// TIA Portal project "uppgift2IndustriellIT" (V18) (continued)
REGION Network 9: if x or y arm is moving for hmi
   RUNG wire#powerrail
      Contact( "InputsDB".Crane.RunArmX )
      { S7_Templates := "SrcType := Int" } NE_Contact(in1 := "Crane Current X Position", in2 := "OutputsDB".CraneOutput.XScalex)
      Coil( "InputsDB".XisMoving )
   END_RUNG
   RUNG wire#powerrail
      Contact( "InputsDB".Crane.RunArmY )
      { S7_Templates := "SrcType := Int" } NE_Contact(in1 := "Crane Current Z Position", in2 := "OutputsDB".CraneOutput.YScalex)
      Coil( "InputsDB".YisMoving )
   END_RUNG
   // the same network as SCL:
   "InputsDB".XisMoving := "InputsDB".Crane.RunArmX AND ("Crane Current X Position" <> "OutputsDB".CraneOutput.XScalex);
   "InputsDB".YisMoving := "InputsDB".Crane.RunArmY AND ("Crane Current Z Position" <> "OutputsDB".CraneOutput.YScalex);
END_REGION
END_FUNCTION

FUNCTION "Outputs" : Void   // FC4, LAD
{ S7_Optimized_Access := 'TRUE' }
VERSION : 0.1
   VAR_TEMP   // added for the SCL form of the ladder/FBD networks
      _w1 : Bool;
      _w2 : Bool;
      _w3 : Bool;
      _w4 : Bool;
   END_VAR
BEGIN

REGION Network 1: Convert MM to raw sensor value which is 27648
   // Calling for example "OutputsDB".CraneOutput.Xmm" with a value from 0-10500mm is going to make the crane move.
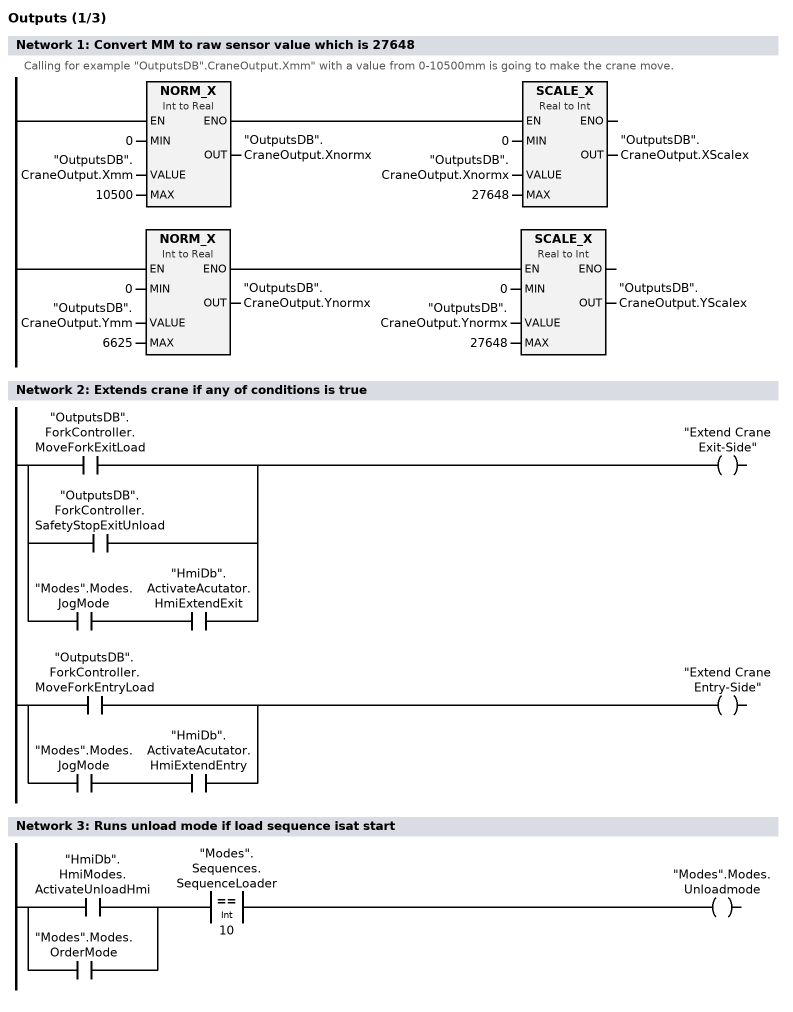
   RUNG wire#powerrail
      { S7_Templates := "[SrcType := Int, DestType := Real]" } Normalize(min := 0, value := "OutputsDB".CraneOutput.Xmm, max := 10500, out => "OutputsDB".CraneOutput.Xnormx)
      { S7_Templates := "[SrcType := Real, DestType := Int]" } Scale(min := 0, value := "OutputsDB".CraneOutput.Xnormx, max := 27648, out => "OutputsDB".CraneOutput.XScalex)
   END_RUNG
   RUNG wire#powerrail
      { S7_Templates := "[SrcType := Int, DestType := Real]" } Normalize(min := 0, value := "OutputsDB".CraneOutput.Ymm, max := 6625, out => "OutputsDB".CraneOutput.Ynormx)
      { S7_Templates := "[SrcType := Real, DestType := Int]" } Scale(min := 0, value := "OutputsDB".CraneOutput.Ynormx, max := 27648, out => "OutputsDB".CraneOutput.YScalex)
   END_RUNG
   // the same network as SCL:
   "OutputsDB".CraneOutput.Xnormx := NORM_X(MIN := 0, VALUE := "OutputsDB".CraneOutput.Xmm, MAX := 10500);
   "OutputsDB".CraneOutput.XScalex := SCALE_X(MIN := 0, VALUE := "OutputsDB".CraneOutput.Xnormx, MAX := 27648);
   "OutputsDB".CraneOutput.Ynormx := NORM_X(MIN := 0, VALUE := "OutputsDB".CraneOutput.Ymm, MAX := 6625);
   "OutputsDB".CraneOutput.YScalex := SCALE_X(MIN := 0, VALUE := "OutputsDB".CraneOutput.Ynormx, MAX := 27648);
END_REGION

REGION Network 2: Extends crane if any of conditions is true
   RUNG wire#powerrail
      Contact( "OutputsDB".ForkController.MoveForkExitLoad )
      wire#w1
      Coil( "Extend Crane Exit-Side" )
   END_RUNG
   RUNG wire#powerrail
      Contact( "OutputsDB".ForkController.SafetyStopExitUnload )
   END_RUNG wire#w1
   RUNG wire#powerrail
      Contact( "Modes".Modes.JogMode )
      Contact( "HmiDb".ActivateAcutator.HmiExtendExit )
   END_RUNG wire#w1
   RUNG wire#powerrail
      Contact( "OutputsDB".ForkController.MoveForkEntryLoad )
      wire#w2
      Coil( "Extend Crane Entry-Side" )
   END_RUNG
   RUNG wire#powerrail
      Contact( "Modes".Modes.JogMode )
      Contact( "HmiDb".ActivateAcutator.HmiExtendEntry )
   END_RUNG wire#w2
   // the same network as SCL:
   "Extend Crane Exit-Side" := "OutputsDB".ForkController.MoveForkExitLoad OR "OutputsDB".ForkController.SafetyStopExitUnload OR ("Modes".Modes.JogMode AND "HmiDb".ActivateAcutator.HmiExtendExit);
   "Extend Crane Entry-Side" := "OutputsDB".ForkController.MoveForkEntryLoad OR ("Modes".Modes.JogMode AND "HmiDb".ActivateAcutator.HmiExtendEntry);
END_REGION

REGION Network 3: Runs unload mode if load sequence isat start
   RUNG wire#powerrail
      Contact( "HmiDb".HmiModes.ActivateUnloadHmi )
      wire#w1
      { S7_Templates := "SrcType := Int" } EQ_Contact(in1 := "Modes".Sequences.SequenceLoader, in2 := 10)
      Coil( "Modes".Modes.Unloadmode )
   END_RUNG
   RUNG wire#powerrail
      Contact( "Modes".Modes.OrderMode )
   END_RUNG wire#w1
   // the same network as SCL:
   "Modes".Modes.Unloadmode := ("HmiDb".HmiModes.ActivateUnloadHmi OR "Modes".Modes.OrderMode) AND ("Modes".Sequences.SequenceLoader = 10);
END_REGION

REGION Network 4: Sets the conveyor speed
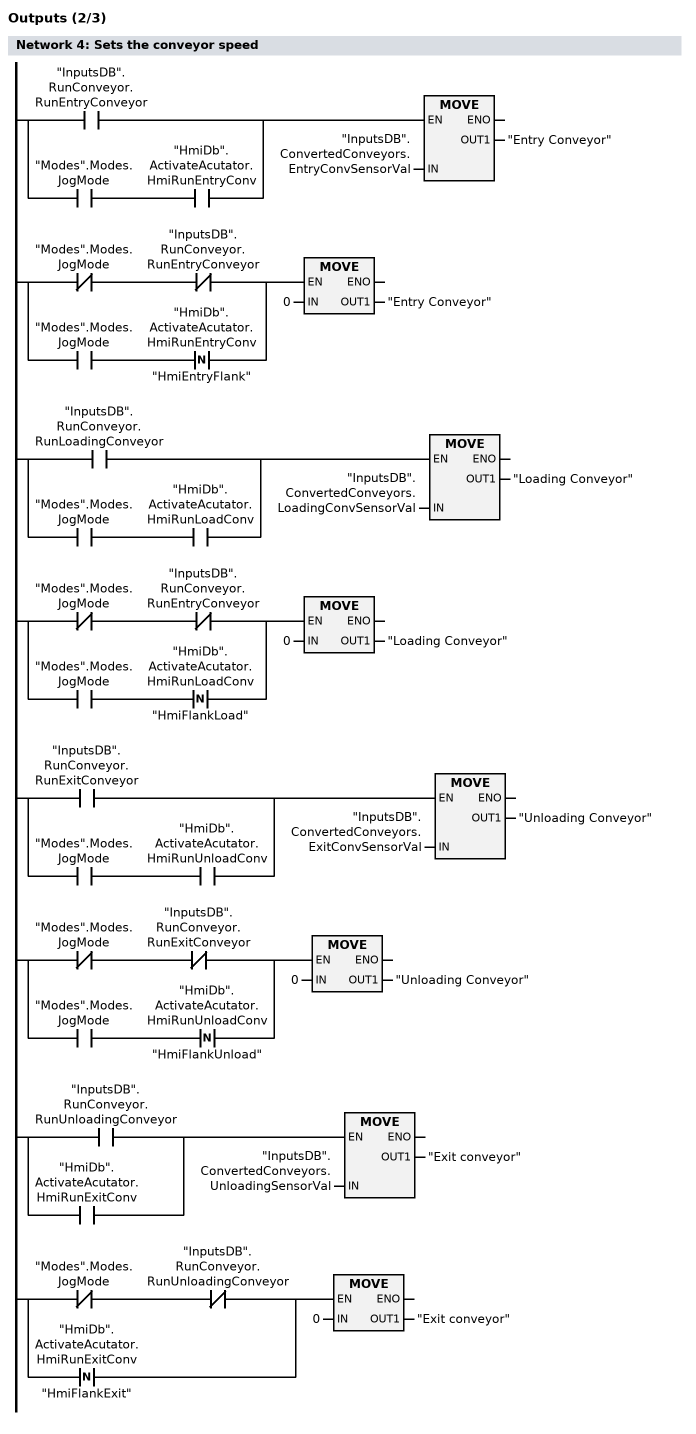
   RUNG wire#powerrail
      Contact( "InputsDB".RunConveyor.RunEntryConveyor )
      wire#w1
      Move(in := "InputsDB".ConvertedConveyors.EntryConvSensorVal, out1 => "Entry Conveyor")
   END_RUNG
   RUNG wire#powerrail
      Contact( "Modes".Modes.JogMode )
      Contact( "HmiDb".ActivateAcutator.HmiRunEntryConv )
   END_RUNG wire#w1
   RUNG wire#powerrail
      I_Contact( "Modes".Modes.JogMode )
      I_Contact( "InputsDB".RunConveyor.RunEntryConveyor )
      wire#w2
      Move(in := 0, out1 => "Entry Conveyor")
   END_RUNG
   RUNG wire#powerrail
      Contact( "Modes".Modes.JogMode )
      N_Contact(operand := "HmiDb".ActivateAcutator.HmiRunEntryConv, bit := "HmiEntryFlank")
   END_RUNG wire#w2
   RUNG wire#powerrail
      Contact( "InputsDB".RunConveyor.RunLoadingConveyor )
      wire#w3
      Move(in := "InputsDB".ConvertedConveyors.LoadingConvSensorVal, out1 => "Loading Conveyor")
   END_RUNG
   RUNG wire#powerrail
      Contact( "Modes".Modes.JogMode )
      Contact( "HmiDb".ActivateAcutator.HmiRunLoadConv )
   END_RUNG wire#w3
   RUNG wire#powerrail
      I_Contact( "Modes".Modes.JogMode )
      I_Contact( "InputsDB".RunConveyor.RunEntryConveyor )
      wire#w4
      Move(in := 0, out1 => "Loading Conveyor")
   END_RUNG
   RUNG wire#powerrail
      Contact( "Modes".Modes.JogMode )
      N_Contact(operand := "HmiDb".ActivateAcutator.HmiRunLoadConv, bit := "HmiFlankLoad")
   END_RUNG wire#w4
   RUNG wire#powerrail
      Contact( "InputsDB".RunConveyor.RunExitConveyor )
      wire#w5
      Move(in := "InputsDB".ConvertedConveyors.ExitConvSensorVal, out1 => "Unloading Conveyor")
   END_RUNG
   RUNG wire#powerrail
      Contact( "Modes".Modes.JogMode )
      Contact( "HmiDb".ActivateAcutator.HmiRunUnloadConv )
   END_RUNG wire#w5
   RUNG wire#powerrail
      I_Contact( "Modes".Modes.JogMode )
      I_Contact( "InputsDB".RunConveyor.RunExitConveyor )
      wire#w6
      Move(in := 0, out1 => "Unloading Conveyor")
   END_RUNG
   RUNG wire#powerrail
      Contact( "Modes".Modes.JogMode )
      N_Contact(operand := "HmiDb".ActivateAcutator.HmiRunUnloadConv, bit := "HmiFlankUnload")
   END_RUNG wire#w6
   RUNG wire#powerrail
      Contact( "InputsDB".RunConveyor.RunUnloadingConveyor )
      wire#w7
      Move(in := "InputsDB".ConvertedConveyors.UnloadingSensorVal, out1 => "Exit conveyor")
   END_RUNG
   RUNG wire#powerrail
      Contact( "HmiDb".ActivateAcutator.HmiRunExitConv )
   END_RUNG wire#w7
   RUNG wire#powerrail
      I_Contact( "Modes".Modes.JogMode )
      I_Contact( "InputsDB".RunConveyor.RunUnloadingConveyor )
      wire#w8
      Move(in := 0, out1 => "Exit conveyor")
   END_RUNG
   RUNG wire#powerrail
      N_Contact(operand := "HmiDb".ActivateAcutator.HmiRunExitConv, bit := "HmiFlankExit")
   END_RUNG wire#w8
   // the same network as SCL:
   IF "InputsDB".RunConveyor.RunEntryConveyor OR ("Modes".Modes.JogMode AND "HmiDb".ActivateAcutator.HmiRunEntryConv) THEN
       "Entry Conveyor" := "InputsDB".ConvertedConveyors.EntryConvSensorVal;
   END_IF;
   #_w1 := "Modes".Modes.JogMode AND NOT "HmiDb".ActivateAcutator.HmiRunEntryConv AND "HmiEntryFlank";   // falling edge of "HmiDb".ActivateAcutator.HmiRunEntryConv
   "HmiEntryFlank" := "HmiDb".ActivateAcutator.HmiRunEntryConv;
   IF (NOT "Modes".Modes.JogMode AND NOT "InputsDB".RunConveyor.RunEntryConveyor) OR #_w1 THEN
       "Entry Conveyor" := 0;
   END_IF;
   IF "InputsDB".RunConveyor.RunLoadingConveyor OR ("Modes".Modes.JogMode AND "HmiDb".ActivateAcutator.HmiRunLoadConv) THEN
       "Loading Conveyor" := "InputsDB".ConvertedConveyors.LoadingConvSensorVal;
   END_IF;
   #_w2 := "Modes".Modes.JogMode AND NOT "HmiDb".ActivateAcutator.HmiRunLoadConv AND "HmiFlankLoad";   // falling edge of "HmiDb".ActivateAcutator.HmiRunLoadConv
   "HmiFlankLoad" := "HmiDb".ActivateAcutator.HmiRunLoadConv;
   IF (NOT "Modes".Modes.JogMode AND NOT "InputsDB".RunConveyor.RunEntryConveyor) OR #_w2 THEN
       "Loading Conveyor" := 0;
   END_IF;
   IF "InputsDB".RunConveyor.RunExitConveyor OR ("Modes".Modes.JogMode AND "HmiDb".ActivateAcutator.HmiRunUnloadConv) THEN
       "Unloading Conveyor" := "InputsDB".ConvertedConveyors.ExitConvSensorVal;
   END_IF;
   #_w3 := "Modes".Modes.JogMode AND NOT "HmiDb".ActivateAcutator.HmiRunUnloadConv AND "HmiFlankUnload";   // falling edge of "HmiDb".ActivateAcutator.HmiRunUnloadConv
   "HmiFlankUnload" := "HmiDb".ActivateAcutator.HmiRunUnloadConv;
   IF (NOT "Modes".Modes.JogMode AND NOT "InputsDB".RunConveyor.RunExitConveyor) OR #_w3 THEN
       "Unloading Conveyor" := 0;
   END_IF;
   IF "InputsDB".RunConveyor.RunUnloadingConveyor OR "HmiDb".ActivateAcutator.HmiRunExitConv THEN
       "Exit conveyor" := "InputsDB".ConvertedConveyors.UnloadingSensorVal;
   END_IF;
   #_w4 := NOT "HmiDb".ActivateAcutator.HmiRunExitConv AND "HmiFlankExit";   // falling edge of "HmiDb".ActivateAcutator.HmiRunExitConv
   "HmiFlankExit" := "HmiDb".ActivateAcutator.HmiRunExitConv;
   IF (NOT "Modes".Modes.JogMode AND NOT "InputsDB".RunConveyor.RunUnloadingConveyor) OR #_w4 THEN
       "Exit conveyor" := 0;
   END_IF;
END_REGION

REGION Network 5: Reset Sequence Resets values on reset has a safety that checks that crane is retracted before moving it
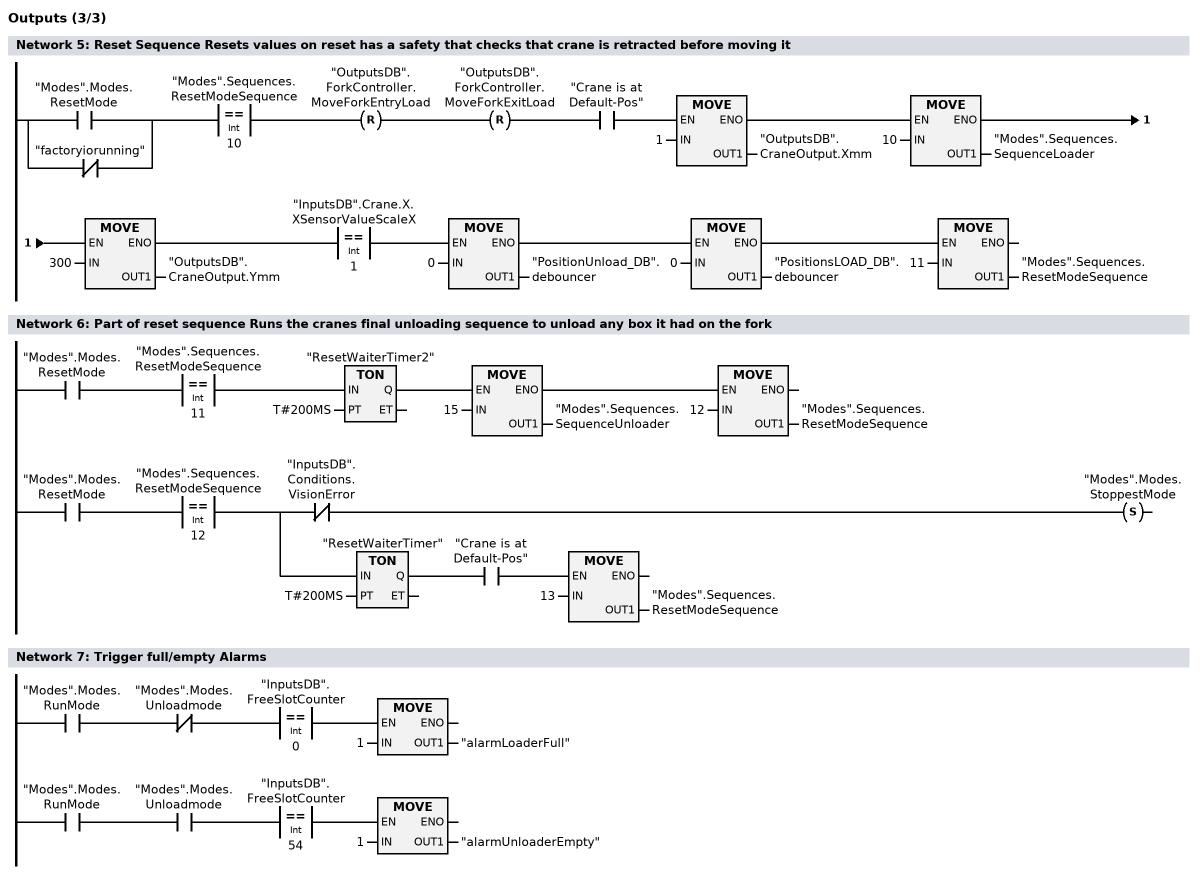
   RUNG wire#powerrail
      Contact( "Modes".Modes.ResetMode )
      wire#w1
      { S7_Templates := "SrcType := Int" } EQ_Contact(in1 := "Modes".Sequences.ResetModeSequence, in2 := 10)
      R_Coil( "OutputsDB".ForkController.MoveForkEntryLoad )
      R_Coil( "OutputsDB".ForkController.MoveForkExitLoad )
      Contact( "Crane is at Default-Pos" )
      Move(in := 1, out1 => "OutputsDB".CraneOutput.Xmm)
      Move(in := 10, out1 => "Modes".Sequences.SequenceLoader)
      Move(in := 300, out1 => "OutputsDB".CraneOutput.Ymm)
      { S7_Templates := "SrcType := Int" } EQ_Contact(in1 := "InputsDB".Crane.X.XSensorValueScaleX, in2 := 1)
      Move(in := 0, out1 => "PositionUnload_DB".debouncer)
      Move(in := 0, out1 => "PositionsLOAD_DB".debouncer)
      Move(in := 11, out1 => "Modes".Sequences.ResetModeSequence)
   END_RUNG
   RUNG wire#powerrail
      I_Contact( "factoryiorunning" )
   END_RUNG wire#w1
   // the same network as SCL:
   #_w1 := ("Modes".Modes.ResetMode OR NOT "factoryiorunning") AND ("Modes".Sequences.ResetModeSequence = 10);
   IF #_w1 THEN
       "OutputsDB".ForkController.MoveForkEntryLoad := FALSE;
       "OutputsDB".ForkController.MoveForkExitLoad := FALSE;
   END_IF;
   #_w2 := #_w1 AND "Crane is at Default-Pos";
   IF #_w2 THEN
       "OutputsDB".CraneOutput.Xmm := 1;
       "Modes".Sequences.SequenceLoader := 10;
       "OutputsDB".CraneOutput.Ymm := 300;
   END_IF;
   IF #_w2 AND ("InputsDB".Crane.X.XSensorValueScaleX = 1) THEN
       "PositionUnload_DB".debouncer := 0;
       "PositionsLOAD_DB".debouncer := 0;
       "Modes".Sequences.ResetModeSequence := 11;
   END_IF;
END_REGION

REGION Network 6: Part of reset sequence Runs the cranes final unloading sequence to unload any box it had on the fork
   "ResetWaiterTimer2".TON(IN := "Modes".Modes.ResetMode AND ("Modes".Sequences.ResetModeSequence = 11),
                           PT := T#200MS);
   IF "ResetWaiterTimer2".Q THEN
       "Modes".Sequences.SequenceUnloader := 15;
       "Modes".Sequences.ResetModeSequence := 12;
   END_IF;
   #_w1 := "Modes".Modes.ResetMode AND ("Modes".Sequences.ResetModeSequence = 12);
   IF #_w1 AND NOT "InputsDB".Conditions.VisionError THEN "Modes".Modes.StoppestMode := TRUE; END_IF;
   "ResetWaiterTimer".TON(IN := #_w1, PT := T#200MS);
   IF "ResetWaiterTimer".Q AND "Crane is at Default-Pos" THEN
       "Modes".Sequences.ResetModeSequence := 13;
   END_IF;
END_REGION

REGION Network 7: Trigger full/empty Alarms
   RUNG wire#powerrail
      Contact( "Modes".Modes.RunMode )
      I_Contact( "Modes".Modes.Unloadmode )
      { S7_Templates := "SrcType := Int" } EQ_Contact(in1 := "InputsDB".FreeSlotCounter, in2 := 0)
      Move(in := 1, out1 => "alarmLoaderFull")
   END_RUNG
   RUNG wire#powerrail
      Contact( "Modes".Modes.RunMode )
      Contact( "Modes".Modes.Unloadmode )
      { S7_Templates := "SrcType := Int" } EQ_Contact(in1 := "InputsDB".FreeSlotCounter, in2 := 54)
      Move(in := 1, out1 => "alarmUnloaderEmpty")
   END_RUNG
   // the same network as SCL:
   IF "Modes".Modes.RunMode AND NOT "Modes".Modes.Unloadmode AND ("InputsDB".FreeSlotCounter = 0) THEN
       "alarmLoaderFull" := 1;
   END_IF;
   IF "Modes".Modes.RunMode AND "Modes".Modes.Unloadmode AND ("InputsDB".FreeSlotCounter = 54) THEN
       "alarmUnloaderEmpty" := 1;
   END_IF;
END_REGION
END_FUNCTION

FUNCTION "ColorDetector" : Void   // FC5, LAD
{ S7_Optimized_Access := 'TRUE' }
VERSION : 0.1
   VAR_TEMP   // added for the SCL form of the ladder/FBD networks
      _w1 : Bool;
      _w2 : Bool;
      _w3 : Bool;
   END_VAR
BEGIN

REGION Network 1: Counts colors
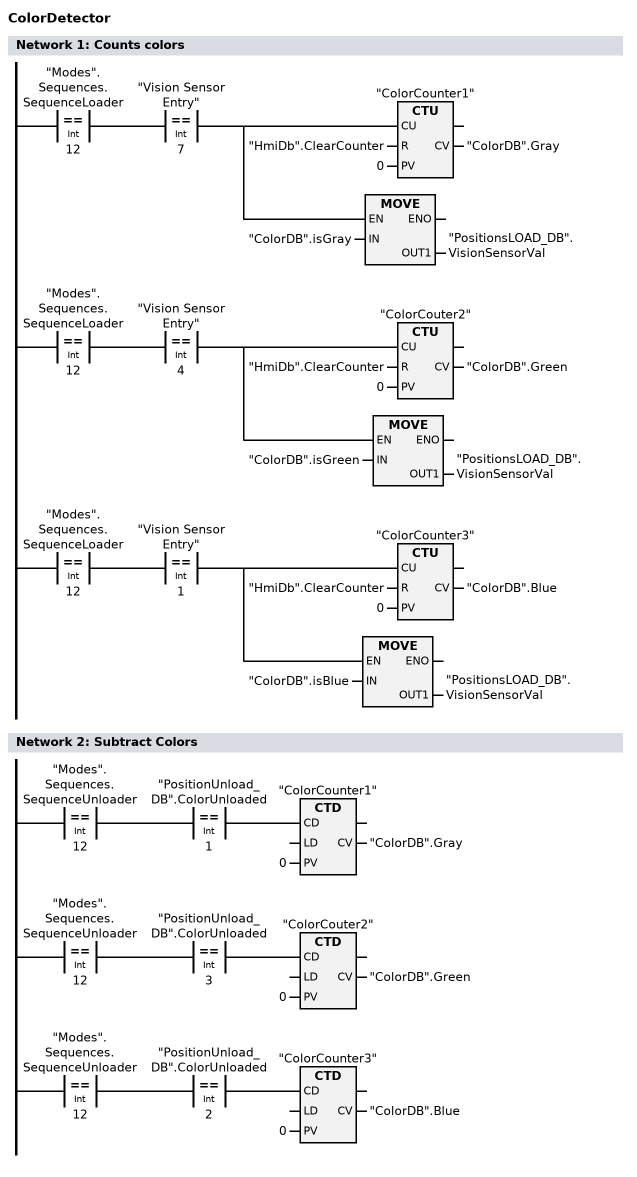
   #_w1 := ("Modes".Sequences.SequenceLoader = 12) AND ("Vision Sensor Entry" = 7);
   "ColorCounter1".CTU(CU := #_w1, R := "HmiDb".ClearCounter, PV := 0, CV => "ColorDB".Gray);
   IF #_w1 THEN "PositionsLOAD_DB".VisionSensorVal := "ColorDB".isGray; END_IF;
   #_w2 := ("Modes".Sequences.SequenceLoader = 12) AND ("Vision Sensor Entry" = 4);
   "ColorCouter2".CTU(CU := #_w2, R := "HmiDb".ClearCounter, PV := 0, CV => "ColorDB".Green);
   IF #_w2 THEN "PositionsLOAD_DB".VisionSensorVal := "ColorDB".isGreen; END_IF;
   #_w3 := ("Modes".Sequences.SequenceLoader = 12) AND ("Vision Sensor Entry" = 1);
   "ColorCounter3".CTU(CU := #_w3, R := "HmiDb".ClearCounter, PV := 0, CV => "ColorDB".Blue);
   IF #_w3 THEN "PositionsLOAD_DB".VisionSensorVal := "ColorDB".isBlue; END_IF;
END_REGION

REGION Network 2: Subtract Colors
   "ColorCounter1".CTD(CD := ("Modes".Sequences.SequenceUnloader = 12) AND ("PositionUnload_DB".ColorUnloaded = 1),
                       PV := 0,
                       CV => "ColorDB".Gray);
   "ColorCouter2".CTD(CD := ("Modes".Sequences.SequenceUnloader = 12) AND ("PositionUnload_DB".ColorUnloaded = 3),
                      PV := 0,
                      CV => "ColorDB".Green);
   "ColorCounter3".CTD(CD := ("Modes".Sequences.SequenceUnloader = 12) AND ("PositionUnload_DB".ColorUnloaded = 2),
                       PV := 0,
                       CV => "ColorDB".Blue);
END_REGION
END_FUNCTION

FUNCTION "SafetyStop" : Void   // FC7, LAD
{ S7_Optimized_Access := 'TRUE' }
VERSION : 0.1
BEGIN

REGION Network 1: Protected stop start
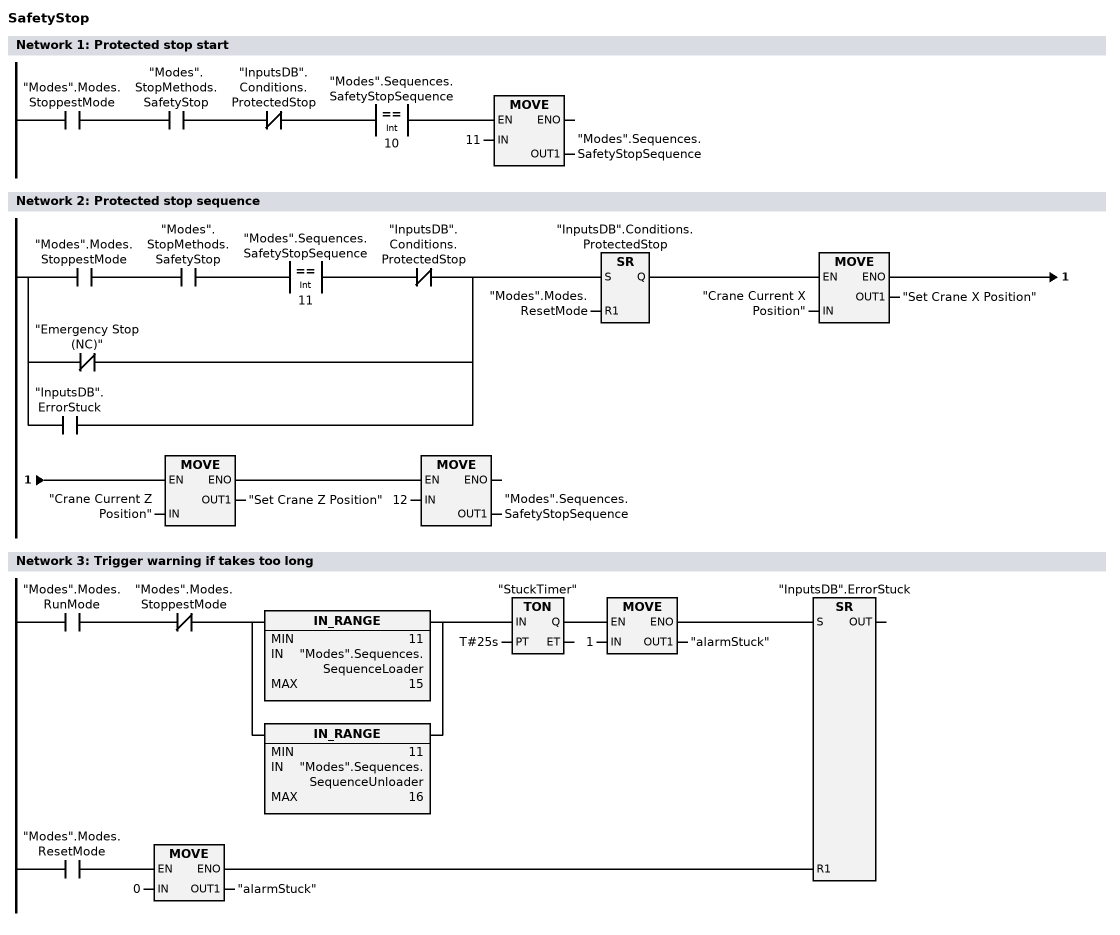
   RUNG wire#powerrail
      Contact( "Modes".Modes.StoppestMode )
      Contact( "Modes".StopMethods.SafetyStop )
      I_Contact( "InputsDB".Conditions.ProtectedStop )
      { S7_Templates := "SrcType := Int" } EQ_Contact(in1 := "Modes".Sequences.SafetyStopSequence, in2 := 10)
      Move(in := 11, out1 => "Modes".Sequences.SafetyStopSequence)
   END_RUNG
   // the same network as SCL:
   IF "Modes".Modes.StoppestMode AND "Modes".StopMethods.SafetyStop AND NOT "InputsDB".Conditions.ProtectedStop AND ("Modes".Sequences.SafetyStopSequence = 10) THEN
       "Modes".Sequences.SafetyStopSequence := 11;
   END_IF;
END_REGION

REGION Network 2: Protected stop sequence
   RUNG wire#powerrail
      Contact( "Modes".Modes.StoppestMode )
      Contact( "Modes".StopMethods.SafetyStop )
      { S7_Templates := "SrcType := Int" } EQ_Contact(in1 := "Modes".Sequences.SafetyStopSequence, in2 := 11)
      I_Contact( "InputsDB".Conditions.ProtectedStop )
      wire#w1
      S_SR(operand := "InputsDB".Conditions.ProtectedStop, r1 := "Modes".Modes.ResetMode)
      Move(in := "Crane Current X Position", out1 => "Set Crane X Position")
      Move(in := "Crane Current Z Position", out1 => "Set Crane Z Position")
      Move(in := 12, out1 => "Modes".Sequences.SafetyStopSequence)
   END_RUNG
   RUNG wire#powerrail
      I_Contact( "Emergency Stop (NC)" )
   END_RUNG wire#w1
   RUNG wire#powerrail
      Contact( "InputsDB".ErrorStuck )
   END_RUNG wire#w1
   // the same network as SCL:
   IF ("Modes".Modes.StoppestMode AND "Modes".StopMethods.SafetyStop AND ("Modes".Sequences.SafetyStopSequence = 11) AND NOT "InputsDB".Conditions.ProtectedStop) OR NOT "Emergency Stop (NC)" OR "InputsDB".ErrorStuck THEN
       "InputsDB".Conditions.ProtectedStop := TRUE;   // SR flip-flop
   END_IF;
   IF "Modes".Modes.ResetMode THEN "InputsDB".Conditions.ProtectedStop := FALSE; END_IF;
   IF "InputsDB".Conditions.ProtectedStop THEN
       "Set Crane X Position" := "Crane Current X Position";
       "Set Crane Z Position" := "Crane Current Z Position";
       "Modes".Sequences.SafetyStopSequence := 12;
   END_IF;
END_REGION

REGION Network 3: Trigger warning if takes too long
   "StuckTimer".TON(IN := "Modes".Modes.RunMode AND NOT "Modes".Modes.StoppestMode AND (((11 <= "Modes".Sequences.SequenceLoader) AND ("Modes".Sequences.SequenceLoader <= 15)) OR ((11 <= "Modes".Sequences.SequenceUnloader) AND ("Modes".Sequences.SequenceUnloader <= 16))),
                    PT := T#25s);
   IF "StuckTimer".Q THEN "alarmStuck" := 1; END_IF;
   IF "Modes".Modes.ResetMode THEN "alarmStuck" := 0; END_IF;
   IF "StuckTimer".Q THEN
       "InputsDB".ErrorStuck := TRUE;   // SR flip-flop
   END_IF;
   IF "Modes".Modes.ResetMode THEN "InputsDB".ErrorStuck := FALSE; END_IF;
END_REGION
END_FUNCTION

(* ===== HMI "HMI_RT_1" =====
system functions are stored by id; their names below are inferred from use
connection "Connection_1": ETHERNET, S7_1500_OMS
connection "HMI_Connection_1": ETHERNET, S7_1500_OMS

